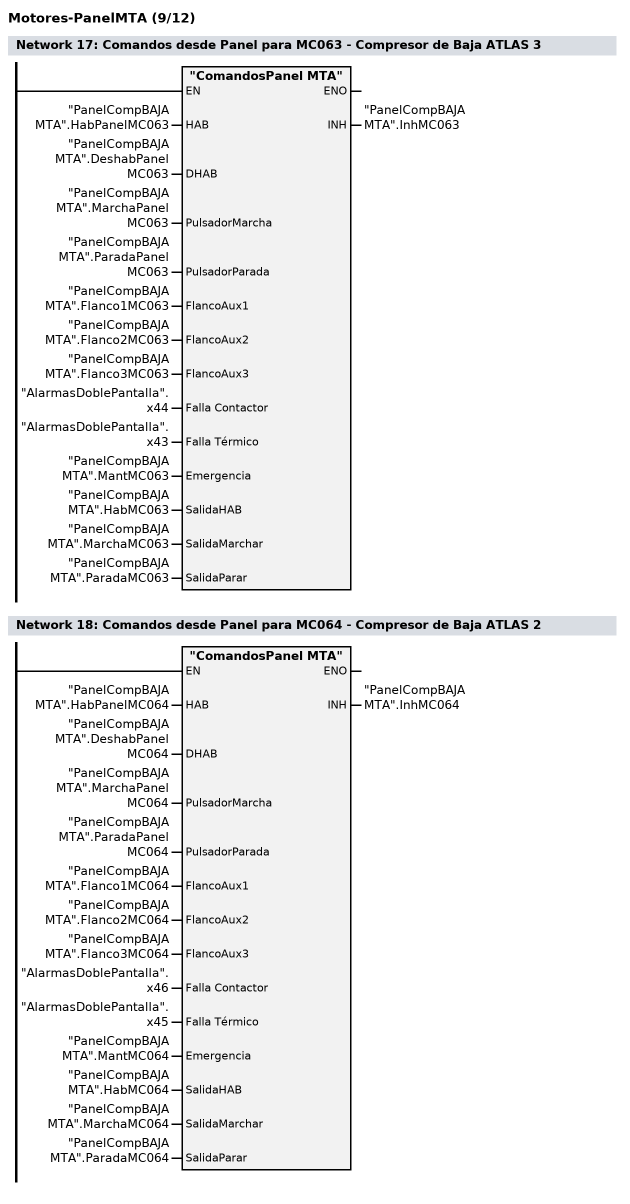
   RUNG wire#powerrail
      "ComandosPanel MTA"(HAB := "PanelCompBAJA MTA".HabPanelMC063, DHAB := "PanelCompBAJA MTA".DeshabPanelMC063, PulsadorMarcha := "PanelCompBAJA MTA".MarchaPanelMC063, PulsadorParada := "PanelCompBAJA MTA".ParadaPanelMC063, FlancoAux1 := "PanelCompBAJA MTA".Flanco1MC063, FlancoAux2 := "PanelCompBAJA MTA".Flanco2MC063, FlancoAux3 := "PanelCompBAJA MTA".Flanco3MC063, "Falla Contactor" := "AlarmasDoblePantalla".x44, "Falla Térmico" := "AlarmasDoblePantalla".x43, Emergencia := "PanelCompBAJA MTA".MantMC063, INH => "PanelCompBAJA MTA".InhMC063, SalidaHAB := "PanelCompBAJA MTA".HabMC063, SalidaMarchar := "PanelCompBAJA MTA".MarchaMC063, SalidaParar := "PanelCompBAJA MTA".ParadaMC063)
   END_RUNG
   // the same network as SCL:
   "ComandosPanel MTA"(HAB := "PanelCompBAJA MTA".HabPanelMC063,
                       DHAB := "PanelCompBAJA MTA".DeshabPanelMC063,
                       PulsadorMarcha := "PanelCompBAJA MTA".MarchaPanelMC063,
                       PulsadorParada := "PanelCompBAJA MTA".ParadaPanelMC063,
                       FlancoAux1 := "PanelCompBAJA MTA".Flanco1MC063,
                       FlancoAux2 := "PanelCompBAJA MTA".Flanco2MC063,
                       FlancoAux3 := "PanelCompBAJA MTA".Flanco3MC063,
                       "Falla Contactor" := "AlarmasDoblePantalla".x44,
                       "Falla Térmico" := "AlarmasDoblePantalla".x43,
                       Emergencia := "PanelCompBAJA MTA".MantMC063,
                       SalidaHAB := "PanelCompBAJA MTA".HabMC063,
                       SalidaMarchar := "PanelCompBAJA MTA".MarchaMC063,
                       SalidaParar := "PanelCompBAJA MTA".ParadaMC063,
                       INH => "PanelCompBAJA MTA".InhMC063);
END_REGION

REGION Network 18: Comandos desde Panel para MC064 - Compresor de Baja ATLAS 2
   RUNG wire#powerrail
      "ComandosPanel MTA"(HAB := "PanelCompBAJA MTA".HabPanelMC064, DHAB := "PanelCompBAJA MTA".DeshabPanelMC064, PulsadorMarcha := "PanelCompBAJA MTA".MarchaPanelMC064, PulsadorParada := "PanelCompBAJA MTA".ParadaPanelMC064, FlancoAux1 := "PanelCompBAJA MTA".Flanco1MC064, FlancoAux2 := "PanelCompBAJA MTA".Flanco2MC064, FlancoAux3 := "PanelCompBAJA MTA".Flanco3MC064, "Falla Contactor" := "AlarmasDoblePantalla".x46, "Falla Térmico" := "AlarmasDoblePantalla".x45, Emergencia := "PanelCompBAJA MTA".MantMC064, INH => "PanelCompBAJA MTA".InhMC064, SalidaHAB := "PanelCompBAJA MTA".HabMC064, SalidaMarchar := "PanelCompBAJA MTA".MarchaMC064, SalidaParar := "PanelCompBAJA MTA".ParadaMC064)
   END_RUNG
   // the same network as SCL:
   "ComandosPanel MTA"(HAB := "PanelCompBAJA MTA".HabPanelMC064,
                       DHAB := "PanelCompBAJA MTA".DeshabPanelMC064,
                       PulsadorMarcha := "PanelCompBAJA MTA".MarchaPanelMC064,
                       PulsadorParada := "PanelCompBAJA MTA".ParadaPanelMC064,
                       FlancoAux1 := "PanelCompBAJA MTA".Flanco1MC064,
                       FlancoAux2 := "PanelCompBAJA MTA".Flanco2MC064,
                       FlancoAux3 := "PanelCompBAJA MTA".Flanco3MC064,
                       "Falla Contactor" := "AlarmasDoblePantalla".x46,
                       "Falla Térmico" := "AlarmasDoblePantalla".x45,
                       Emergencia := "PanelCompBAJA MTA".MantMC064,
                       SalidaHAB := "PanelCompBAJA MTA".HabMC064,
                       SalidaMarchar := "PanelCompBAJA MTA".MarchaMC064,
                       SalidaParar := "PanelCompBAJA MTA".ParadaMC064,
                       INH => "PanelCompBAJA MTA".InhMC064);
END_REGION

REGION Network 19: Comandos desde Panel para MS050 - Secador de Alta ABC1
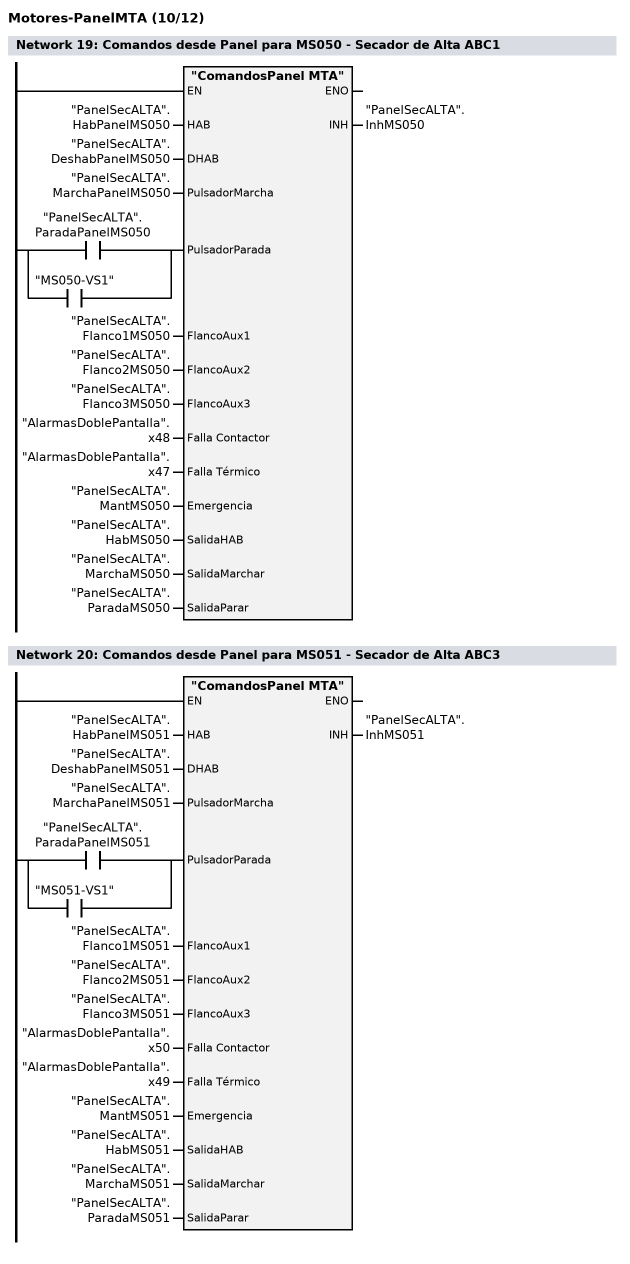
   RUNG wire#powerrail
      "ComandosPanel MTA"(HAB := "PanelSecALTA".HabPanelMS050, DHAB := "PanelSecALTA".DeshabPanelMS050, PulsadorMarcha := "PanelSecALTA".MarchaPanelMS050, PulsadorParada := wire#w1, FlancoAux1 := "PanelSecALTA".Flanco1MS050, FlancoAux2 := "PanelSecALTA".Flanco2MS050, FlancoAux3 := "PanelSecALTA".Flanco3MS050, "Falla Contactor" := "AlarmasDoblePantalla".x48, "Falla Térmico" := "AlarmasDoblePantalla".x47, Emergencia := "PanelSecALTA".MantMS050, INH => "PanelSecALTA".InhMS050, SalidaHAB := "PanelSecALTA".HabMS050, SalidaMarchar := "PanelSecALTA".MarchaMS050, SalidaParar := "PanelSecALTA".ParadaMS050)
   END_RUNG
   RUNG wire#powerrail
      Contact( "PanelSecALTA".ParadaPanelMS050 )
   END_RUNG wire#w1
   RUNG wire#powerrail
      Contact( "MS050-VS1" )
   END_RUNG wire#w1
   // the same network as SCL:
   "ComandosPanel MTA"(HAB := "PanelSecALTA".HabPanelMS050,
                       DHAB := "PanelSecALTA".DeshabPanelMS050,
                       PulsadorMarcha := "PanelSecALTA".MarchaPanelMS050,
                       PulsadorParada := "PanelSecALTA".ParadaPanelMS050 OR "MS050-VS1",
                       FlancoAux1 := "PanelSecALTA".Flanco1MS050,
                       FlancoAux2 := "PanelSecALTA".Flanco2MS050,
                       FlancoAux3 := "PanelSecALTA".Flanco3MS050,
                       "Falla Contactor" := "AlarmasDoblePantalla".x48,
                       "Falla Térmico" := "AlarmasDoblePantalla".x47,
                       Emergencia := "PanelSecALTA".MantMS050,
                       SalidaHAB := "PanelSecALTA".HabMS050,
                       SalidaMarchar := "PanelSecALTA".MarchaMS050,
                       SalidaParar := "PanelSecALTA".ParadaMS050,
                       INH => "PanelSecALTA".InhMS050);
END_REGION

REGION Network 20: Comandos desde Panel para MS051 - Secador de Alta ABC3
   RUNG wire#powerrail
      "ComandosPanel MTA"(HAB := "PanelSecALTA".HabPanelMS051, DHAB := "PanelSecALTA".DeshabPanelMS051, PulsadorMarcha := "PanelSecALTA".MarchaPanelMS051, PulsadorParada := wire#w1, FlancoAux1 := "PanelSecALTA".Flanco1MS051, FlancoAux2 := "PanelSecALTA".Flanco2MS051, FlancoAux3 := "PanelSecALTA".Flanco3MS051, "Falla Contactor" := "AlarmasDoblePantalla".x50, "Falla Térmico" := "AlarmasDoblePantalla".x49, Emergencia := "PanelSecALTA".MantMS051, INH => "PanelSecALTA".InhMS051, SalidaHAB := "PanelSecALTA".HabMS051, SalidaMarchar := "PanelSecALTA".MarchaMS051, SalidaParar := "PanelSecALTA".ParadaMS051)
   END_RUNG
   RUNG wire#powerrail
      Contact( "PanelSecALTA".ParadaPanelMS051 )
   END_RUNG wire#w1
   RUNG wire#powerrail
      Contact( "MS051-VS1" )
   END_RUNG wire#w1
   // the same network as SCL:
   "ComandosPanel MTA"(HAB := "PanelSecALTA".HabPanelMS051,
                       DHAB := "PanelSecALTA".DeshabPanelMS051,
                       PulsadorMarcha := "PanelSecALTA".MarchaPanelMS051,
                       PulsadorParada := "PanelSecALTA".ParadaPanelMS051 OR "MS051-VS1",
                       FlancoAux1 := "PanelSecALTA".Flanco1MS051,
                       FlancoAux2 := "PanelSecALTA".Flanco2MS051,
                       FlancoAux3 := "PanelSecALTA".Flanco3MS051,
                       "Falla Contactor" := "AlarmasDoblePantalla".x50,
                       "Falla Térmico" := "AlarmasDoblePantalla".x49,
                       Emergencia := "PanelSecALTA".MantMS051,
                       SalidaHAB := "PanelSecALTA".HabMS051,
                       SalidaMarchar := "PanelSecALTA".MarchaMS051,
                       SalidaParar := "PanelSecALTA".ParadaMS051,
                       INH => "PanelSecALTA".InhMS051);
END_REGION

REGION Network 21: Comandos desde Panel para MS052 - Secador de Alta ABC2
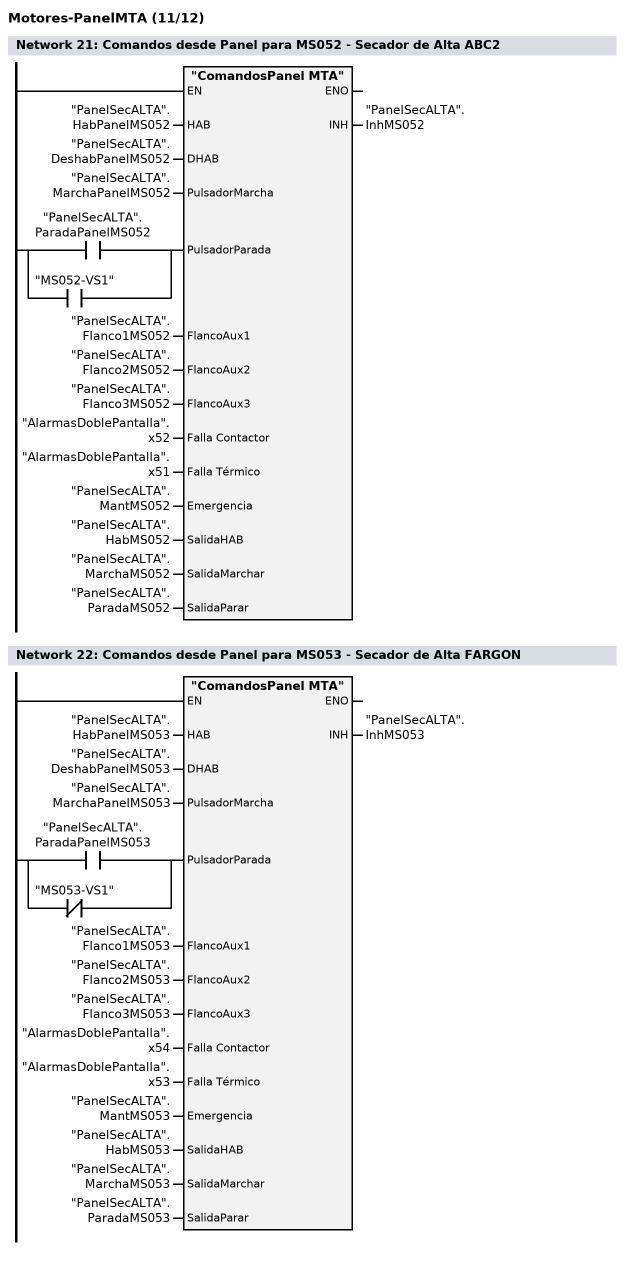
   RUNG wire#powerrail
      "ComandosPanel MTA"(HAB := "PanelSecALTA".HabPanelMS052, DHAB := "PanelSecALTA".DeshabPanelMS052, PulsadorMarcha := "PanelSecALTA".MarchaPanelMS052, PulsadorParada := wire#w1, FlancoAux1 := "PanelSecALTA".Flanco1MS052, FlancoAux2 := "PanelSecALTA".Flanco2MS052, FlancoAux3 := "PanelSecALTA".Flanco3MS052, "Falla Contactor" := "AlarmasDoblePantalla".x52, "Falla Térmico" := "AlarmasDoblePantalla".x51, Emergencia := "PanelSecALTA".MantMS052, INH => "PanelSecALTA".InhMS052, SalidaHAB := "PanelSecALTA".HabMS052, SalidaMarchar := "PanelSecALTA".MarchaMS052, SalidaParar := "PanelSecALTA".ParadaMS052)
   END_RUNG
   RUNG wire#powerrail
      Contact( "PanelSecALTA".ParadaPanelMS052 )
   END_RUNG wire#w1
   RUNG wire#powerrail
      Contact( "MS052-VS1" )
   END_RUNG wire#w1
   // the same network as SCL:
   "ComandosPanel MTA"(HAB := "PanelSecALTA".HabPanelMS052,
                       DHAB := "PanelSecALTA".DeshabPanelMS052,
                       PulsadorMarcha := "PanelSecALTA".MarchaPanelMS052,
                       PulsadorParada := "PanelSecALTA".ParadaPanelMS052 OR "MS052-VS1",
                       FlancoAux1 := "PanelSecALTA".Flanco1MS052,
                       FlancoAux2 := "PanelSecALTA".Flanco2MS052,
                       FlancoAux3 := "PanelSecALTA".Flanco3MS052,
                       "Falla Contactor" := "AlarmasDoblePantalla".x52,
                       "Falla Térmico" := "AlarmasDoblePantalla".x51,
                       Emergencia := "PanelSecALTA".MantMS052,
                       SalidaHAB := "PanelSecALTA".HabMS052,
                       SalidaMarchar := "PanelSecALTA".MarchaMS052,
                       SalidaParar := "PanelSecALTA".ParadaMS052,
                       INH => "PanelSecALTA".InhMS052);
END_REGION

REGION Network 22: Comandos desde Panel para MS053 - Secador de Alta FARGON
   RUNG wire#powerrail
      "ComandosPanel MTA"(HAB := "PanelSecALTA".HabPanelMS053, DHAB := "PanelSecALTA".DeshabPanelMS053, PulsadorMarcha := "PanelSecALTA".MarchaPanelMS053, PulsadorParada := wire#w1, FlancoAux1 := "PanelSecALTA".Flanco1MS053, FlancoAux2 := "PanelSecALTA".Flanco2MS053, FlancoAux3 := "PanelSecALTA".Flanco3MS053, "Falla Contactor" := "AlarmasDoblePantalla".x54, "Falla Térmico" := "AlarmasDoblePantalla".x53, Emergencia := "PanelSecALTA".MantMS053, INH => "PanelSecALTA".InhMS053, SalidaHAB := "PanelSecALTA".HabMS053, SalidaMarchar := "PanelSecALTA".MarchaMS053, SalidaParar := "PanelSecALTA".ParadaMS053)
   END_RUNG
   RUNG wire#powerrail
      Contact( "PanelSecALTA".ParadaPanelMS053 )
   END_RUNG wire#w1
   RUNG wire#powerrail
      I_Contact( "MS053-VS1" )
   END_RUNG wire#w1
   // the same network as SCL:
   "ComandosPanel MTA"(HAB := "PanelSecALTA".HabPanelMS053,
                       DHAB := "PanelSecALTA".DeshabPanelMS053,
                       PulsadorMarcha := "PanelSecALTA".MarchaPanelMS053,
                       PulsadorParada := "PanelSecALTA".ParadaPanelMS053 OR NOT "MS053-VS1",
                       FlancoAux1 := "PanelSecALTA".Flanco1MS053,
                       FlancoAux2 := "PanelSecALTA".Flanco2MS053,
                       FlancoAux3 := "PanelSecALTA".Flanco3MS053,
                       "Falla Contactor" := "AlarmasDoblePantalla".x54,
                       "Falla Térmico" := "AlarmasDoblePantalla".x53,
                       Emergencia := "PanelSecALTA".MantMS053,
                       SalidaHAB := "PanelSecALTA".HabMS053,
                       SalidaMarchar := "PanelSecALTA".MarchaMS053,
                       SalidaParar := "PanelSecALTA".ParadaMS053,
                       INH => "PanelSecALTA".InhMS053);
END_REGION

REGION Network 23: Comandos desde Panel para MS054 - Secador de Baja SULLAIR 1
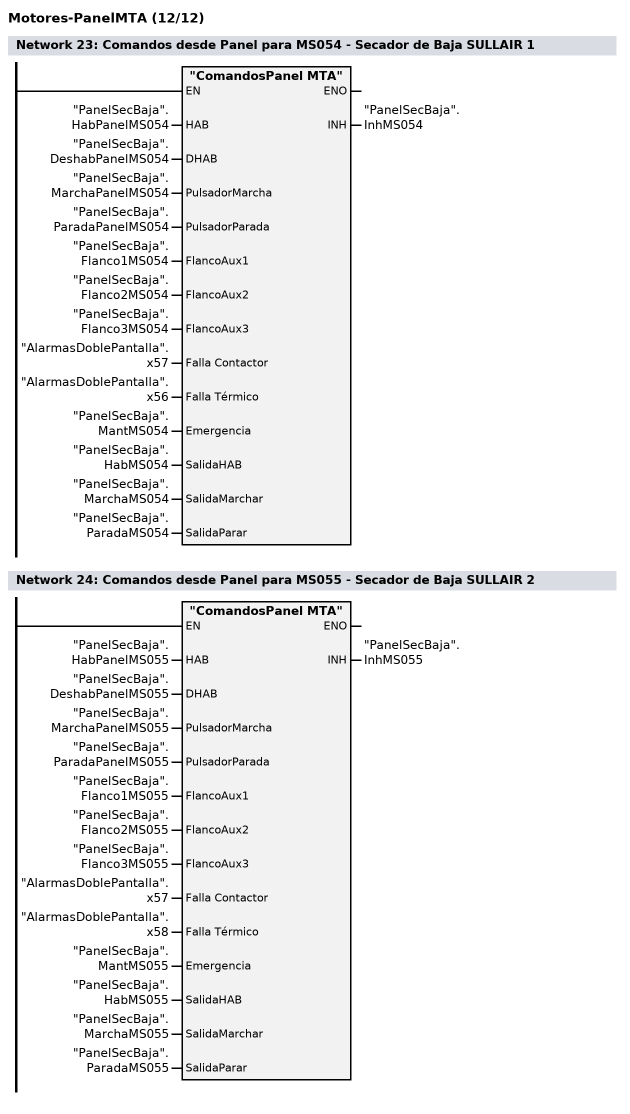
   RUNG wire#powerrail
      "ComandosPanel MTA"(HAB := "PanelSecBaja".HabPanelMS054, DHAB := "PanelSecBaja".DeshabPanelMS054, PulsadorMarcha := "PanelSecBaja".MarchaPanelMS054, PulsadorParada := "PanelSecBaja".ParadaPanelMS054, FlancoAux1 := "PanelSecBaja".Flanco1MS054, FlancoAux2 := "PanelSecBaja".Flanco2MS054, FlancoAux3 := "PanelSecBaja".Flanco3MS054, "Falla Contactor" := "AlarmasDoblePantalla".x57, "Falla Térmico" := "AlarmasDoblePantalla".x56, Emergencia := "PanelSecBaja".MantMS054, INH => "PanelSecBaja".InhMS054, SalidaHAB := "PanelSecBaja".HabMS054, SalidaMarchar := "PanelSecBaja".MarchaMS054, SalidaParar := "PanelSecBaja".ParadaMS054)
   END_RUNG
   // the same network as SCL:
   "ComandosPanel MTA"(HAB := "PanelSecBaja".HabPanelMS054,
                       DHAB := "PanelSecBaja".DeshabPanelMS054,
                       PulsadorMarcha := "PanelSecBaja".MarchaPanelMS054,
                       PulsadorParada := "PanelSecBaja".ParadaPanelMS054,
                       FlancoAux1 := "PanelSecBaja".Flanco1MS054,
                       FlancoAux2 := "PanelSecBaja".Flanco2MS054,
                       FlancoAux3 := "PanelSecBaja".Flanco3MS054,
                       "Falla Contactor" := "AlarmasDoblePantalla".x57,
                       "Falla Térmico" := "AlarmasDoblePantalla".x56,
                       Emergencia := "PanelSecBaja".MantMS054,
                       SalidaHAB := "PanelSecBaja".HabMS054,
                       SalidaMarchar := "PanelSecBaja".MarchaMS054,
                       SalidaParar := "PanelSecBaja".ParadaMS054,
                       INH => "PanelSecBaja".InhMS054);
END_REGION

REGION Network 24: Comandos desde Panel para MS055 - Secador de Baja SULLAIR 2
   RUNG wire#powerrail
      "ComandosPanel MTA"(HAB := "PanelSecBaja".HabPanelMS055, DHAB := "PanelSecBaja".DeshabPanelMS055, PulsadorMarcha := "PanelSecBaja".MarchaPanelMS055, PulsadorParada := "PanelSecBaja".ParadaPanelMS055, FlancoAux1 := "PanelSecBaja".Flanco1MS055, FlancoAux2 := "PanelSecBaja".Flanco2MS055, FlancoAux3 := "PanelSecBaja".Flanco3MS055, "Falla Contactor" := "AlarmasDoblePantalla".x57, "Falla Térmico" := "AlarmasDoblePantalla".x58, Emergencia := "PanelSecBaja".MantMS055, INH => "PanelSecBaja".InhMS055, SalidaHAB := "PanelSecBaja".HabMS055, SalidaMarchar := "PanelSecBaja".MarchaMS055, SalidaParar := "PanelSecBaja".ParadaMS055)
   END_RUNG
   // the same network as SCL:
   "ComandosPanel MTA"(HAB := "PanelSecBaja".HabPanelMS055,
                       DHAB := "PanelSecBaja".DeshabPanelMS055,
                       PulsadorMarcha := "PanelSecBaja".MarchaPanelMS055,
                       PulsadorParada := "PanelSecBaja".ParadaPanelMS055,
                       FlancoAux1 := "PanelSecBaja".Flanco1MS055,
                       FlancoAux2 := "PanelSecBaja".Flanco2MS055,
                       FlancoAux3 := "PanelSecBaja".Flanco3MS055,
                       "Falla Contactor" := "AlarmasDoblePantalla".x57,
                       "Falla Térmico" := "AlarmasDoblePantalla".x58,
                       Emergencia := "PanelSecBaja".MantMS055,
                       SalidaHAB := "PanelSecBaja".HabMS055,
                       SalidaMarchar := "PanelSecBaja".MarchaMS055,
                       SalidaParar := "PanelSecBaja".ParadaMS055,
                       INH => "PanelSecBaja".InhMS055);
END_REGION
END_FUNCTION

FUNCTION "ComandosPanel MTA" : Void   // FC19, LAD
{ S7_Optimized_Access := 'FALSE' }
VERSION : 0.1
   VAR_TEMP   // added for the SCL form of the ladder/FBD networks
      _w1 : Bool;
   END_VAR
BEGIN

REGION Network 1
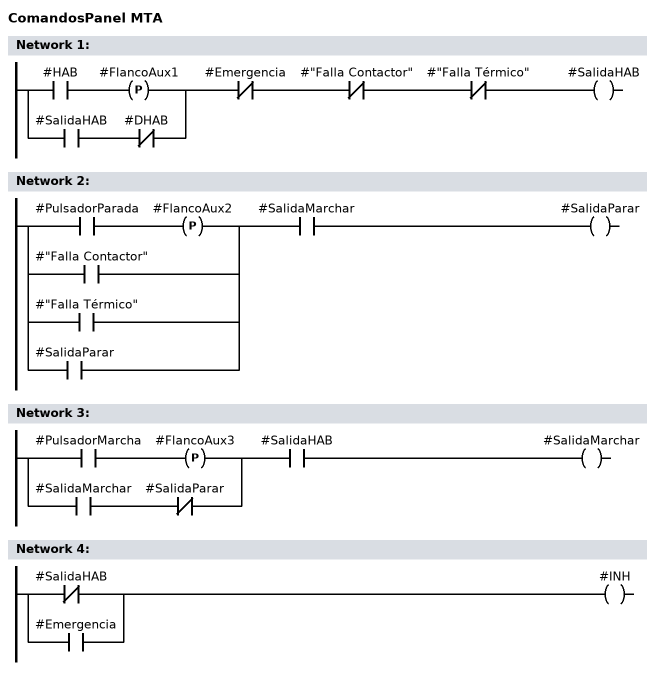
   RUNG wire#powerrail
      Contact( #HAB )
      P_Trig( #FlancoAux1 )
      wire#w1
      I_Contact( #Emergencia )
      I_Contact( #"Falla Contactor" )
      I_Contact( #"Falla Térmico" )
      Coil( #SalidaHAB )
   END_RUNG
   RUNG wire#powerrail
      Contact( #SalidaHAB )
      I_Contact( #DHAB )
   END_RUNG wire#w1
   // the same network as SCL:
   #_w1 := #HAB AND NOT #FlancoAux1;   // rising edge
   #FlancoAux1 := #HAB;
   #SalidaHAB := (#_w1 OR (#SalidaHAB AND NOT #DHAB)) AND NOT #Emergencia AND NOT #"Falla Contactor" AND NOT #"Falla Térmico";
END_REGION

REGION Network 2
   RUNG wire#powerrail
      Contact( #PulsadorParada )
      P_Trig( #FlancoAux2 )
      wire#w1
      Contact( #SalidaMarchar )
      Coil( #SalidaParar )
   END_RUNG
   RUNG wire#powerrail
      Contact( #"Falla Contactor" )
   END_RUNG wire#w1
   RUNG wire#powerrail
      Contact( #"Falla Térmico" )
   END_RUNG wire#w1
   RUNG wire#powerrail
      Contact( #SalidaParar )
   END_RUNG wire#w1
   // the same network as SCL:
   #_w1 := #PulsadorParada AND NOT #FlancoAux2;   // rising edge
   #FlancoAux2 := #PulsadorParada;
   #SalidaParar := (#_w1 OR #"Falla Contactor" OR #"Falla Térmico" OR #SalidaParar) AND #SalidaMarchar;
END_REGION

REGION Network 3
   RUNG wire#powerrail
      Contact( #PulsadorMarcha )
      P_Trig( #FlancoAux3 )
      wire#w1
      Contact( #SalidaHAB )
      Coil( #SalidaMarchar )
   END_RUNG
   RUNG wire#powerrail
      Contact( #SalidaMarchar )
      I_Contact( #SalidaParar )
   END_RUNG wire#w1
   // the same network as SCL:
   #_w1 := #PulsadorMarcha AND NOT #FlancoAux3;   // rising edge
   #FlancoAux3 := #PulsadorMarcha;
   #SalidaMarchar := (#_w1 OR (#SalidaMarchar AND NOT #SalidaParar)) AND #SalidaHAB;
END_REGION

REGION Network 4
   RUNG wire#powerrail
      I_Contact( #SalidaHAB )
      wire#w1
      Coil( #INH )
   END_RUNG
   RUNG wire#powerrail
      Contact( #Emergencia )
   END_RUNG wire#w1
   // the same network as SCL:
   #INH := NOT #SalidaHAB OR #Emergencia;
END_REGION
END_FUNCTION

FUNCTION "FC-ANIM-CMP" : Void   // FC43, LAD
{ S7_Optimized_Access := 'FALSE' }
VERSION : 0.1
BEGIN

REGION Network 1
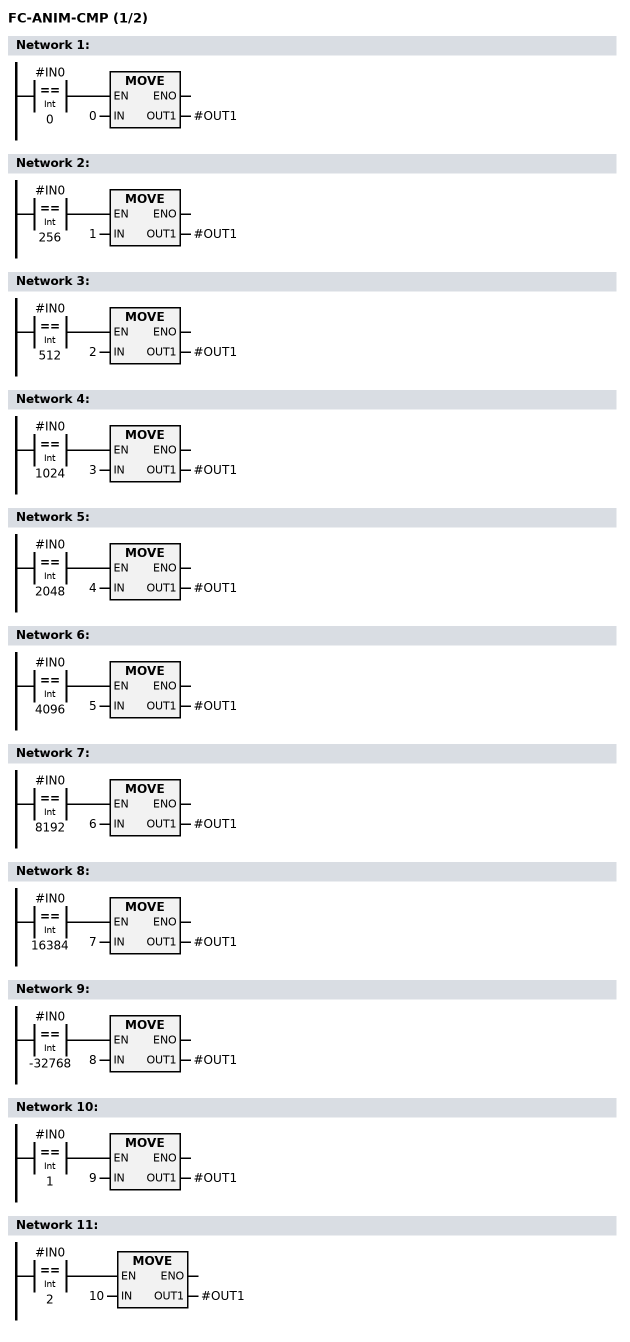
   RUNG wire#powerrail
      { S7_Templates := "SrcType := Int" } EQ_Contact(in1 := #IN0, in2 := 0)
      { S7_GenerateENO := "TRUE" } Move(in := 0, out1 => #OUT1)
   END_RUNG
   // the same network as SCL:
   IF #IN0 = 0 THEN #OUT1 := 0; END_IF;
END_REGION

REGION Network 2
   RUNG wire#powerrail
      { S7_Templates := "SrcType := Int" } EQ_Contact(in1 := #IN0, in2 := 256)
      { S7_GenerateENO := "TRUE" } Move(in := 1, out1 => #OUT1)
   END_RUNG
   // the same network as SCL:
   IF #IN0 = 256 THEN #OUT1 := 1; END_IF;
END_REGION

REGION Network 3
   RUNG wire#powerrail
      { S7_Templates := "SrcType := Int" } EQ_Contact(in1 := #IN0, in2 := 512)
      { S7_GenerateENO := "TRUE" } Move(in := 2, out1 => #OUT1)
   END_RUNG
   // the same network as SCL:
   IF #IN0 = 512 THEN #OUT1 := 2; END_IF;
END_REGION

REGION Network 4
   RUNG wire#powerrail
      { S7_Templates := "SrcType := Int" } EQ_Contact(in1 := #IN0, in2 := 1024)
      { S7_GenerateENO := "TRUE" } Move(in := 3, out1 => #OUT1)
   END_RUNG
   // the same network as SCL:
   IF #IN0 = 1024 THEN #OUT1 := 3; END_IF;
END_REGION

REGION Network 5
   RUNG wire#powerrail
      { S7_Templates := "SrcType := Int" } EQ_Contact(in1 := #IN0, in2 := 2048)
      { S7_GenerateENO := "TRUE" } Move(in := 4, out1 => #OUT1)
   END_RUNG
   // the same network as SCL:
   IF #IN0 = 2048 THEN #OUT1 := 4; END_IF;
END_REGION

REGION Network 6
   RUNG wire#powerrail
      { S7_Templates := "SrcType := Int" } EQ_Contact(in1 := #IN0, in2 := 4096)
      { S7_GenerateENO := "TRUE" } Move(in := 5, out1 => #OUT1)
   END_RUNG
   // the same network as SCL:
   IF #IN0 = 4096 THEN #OUT1 := 5; END_IF;
END_REGION

REGION Network 7
   RUNG wire#powerrail
      { S7_Templates := "SrcType := Int" } EQ_Contact(in1 := #IN0, in2 := 8192)
      { S7_GenerateENO := "TRUE" } Move(in := 6, out1 => #OUT1)
   END_RUNG
   // the same network as SCL:
   IF #IN0 = 8192 THEN #OUT1 := 6; END_IF;
END_REGION

REGION Network 8
   RUNG wire#powerrail
      { S7_Templates := "SrcType := Int" } EQ_Contact(in1 := #IN0, in2 := 16384)
      { S7_GenerateENO := "TRUE" } Move(in := 7, out1 => #OUT1)
   END_RUNG
   // the same network as SCL:
   IF #IN0 = 16384 THEN #OUT1 := 7; END_IF;
END_REGION

REGION Network 9
   RUNG wire#powerrail
      { S7_Templates := "SrcType := Int" } EQ_Contact(in1 := #IN0, in2 := -32768)
      { S7_GenerateENO := "TRUE" } Move(in := 8, out1 => #OUT1)
   END_RUNG
   // the same network as SCL:
   IF #IN0 = (-32768) THEN #OUT1 := 8; END_IF;
END_REGION

REGION Network 10
   RUNG wire#powerrail
      { S7_Templates := "SrcType := Int" } EQ_Contact(in1 := #IN0, in2 := 1)
      { S7_GenerateENO := "TRUE" } Move(in := 9, out1 => #OUT1)
   END_RUNG
   // the same network as SCL:
   IF #IN0 = 1 THEN #OUT1 := 9; END_IF;
END_REGION

REGION Network 11
   RUNG wire#powerrail
      { S7_Templates := "SrcType := Int" } EQ_Contact(in1 := #IN0, in2 := 2)
      { S7_GenerateENO := "TRUE" } Move(in := 10, out1 => #OUT1)
   END_RUNG
   // the same network as SCL:
   IF #IN0 = 2 THEN #OUT1 := 10; END_IF;
END_REGION

REGION Network 12
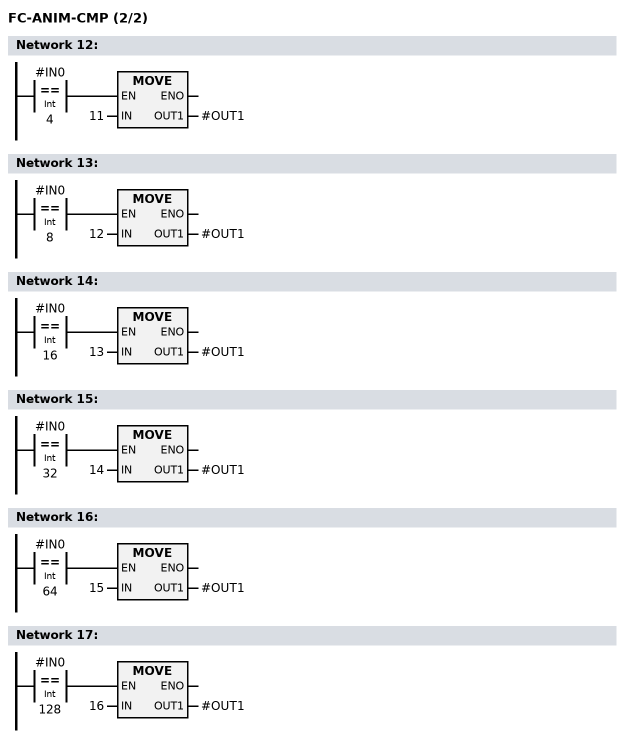
   RUNG wire#powerrail
      { S7_Templates := "SrcType := Int" } EQ_Contact(in1 := #IN0, in2 := 4)
      { S7_GenerateENO := "TRUE" } Move(in := 11, out1 => #OUT1)
   END_RUNG
   // the same network as SCL:
   IF #IN0 = 4 THEN #OUT1 := 11; END_IF;
END_REGION

REGION Network 13
   RUNG wire#powerrail
      { S7_Templates := "SrcType := Int" } EQ_Contact(in1 := #IN0, in2 := 8)
      { S7_GenerateENO := "TRUE" } Move(in := 12, out1 => #OUT1)
   END_RUNG
   // the same network as SCL:
   IF #IN0 = 8 THEN #OUT1 := 12; END_IF;
END_REGION

REGION Network 14
   RUNG wire#powerrail
      { S7_Templates := "SrcType := Int" } EQ_Contact(in1 := #IN0, in2 := 16)
      { S7_GenerateENO := "TRUE" } Move(in := 13, out1 => #OUT1)
   END_RUNG
   // the same network as SCL:
   IF #IN0 = 16 THEN #OUT1 := 13; END_IF;
END_REGION

REGION Network 15
   RUNG wire#powerrail
      { S7_Templates := "SrcType := Int" } EQ_Contact(in1 := #IN0, in2 := 32)
      { S7_GenerateENO := "TRUE" } Move(in := 14, out1 => #OUT1)
   END_RUNG
   // the same network as SCL:
   IF #IN0 = 32 THEN #OUT1 := 14; END_IF;
END_REGION

REGION Network 16
   RUNG wire#powerrail
      { S7_Templates := "SrcType := Int" } EQ_Contact(in1 := #IN0, in2 := 64)
      { S7_GenerateENO := "TRUE" } Move(in := 15, out1 => #OUT1)
   END_RUNG
   // the same network as SCL:
   IF #IN0 = 64 THEN #OUT1 := 15; END_IF;
END_REGION

REGION Network 17
   RUNG wire#powerrail
      { S7_Templates := "SrcType := Int" } EQ_Contact(in1 := #IN0, in2 := 128)
      { S7_GenerateENO := "TRUE" } Move(in := 16, out1 => #OUT1)
   END_RUNG
   // the same network as SCL:
   IF #IN0 = 128 THEN #OUT1 := 16; END_IF;
END_REGION
END_FUNCTION

// folder: Panel/Iluminación

FUNCTION "IluminaciónMTA" : Void   // FC23, LAD
{ S7_Optimized_Access := 'FALSE' }
VERSION : 0.1
// LUC - 05/08/2020
   VAR_TEMP   // added for the SCL form of the ladder/FBD networks
      _s5time1 : S5Time;
   END_VAR
BEGIN

REGION Network 1: Seteo de temporizador desde panel
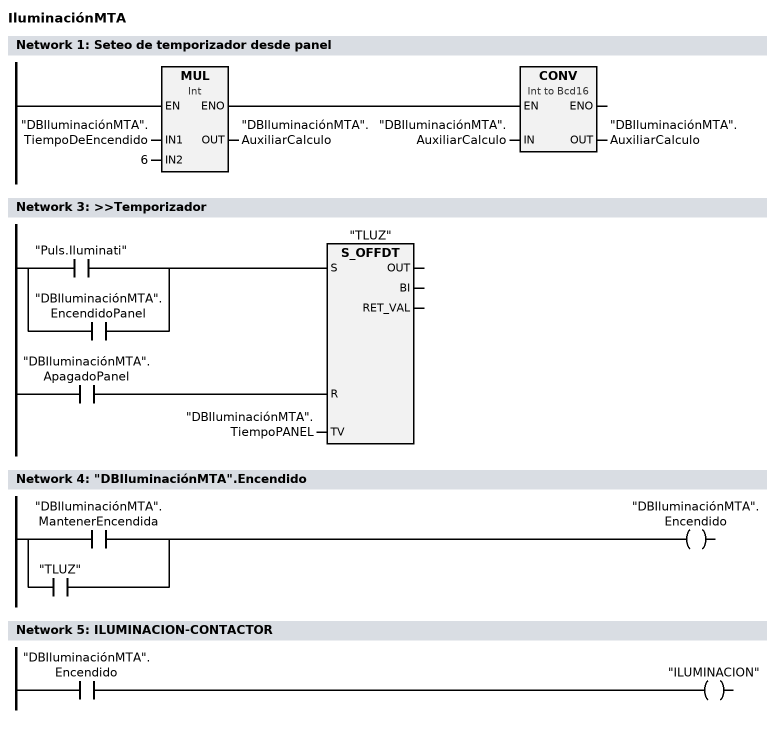
   RUNG wire#powerrail
      { S7_Templates := "SrcType := Int"; S7_GenerateENO := "TRUE" } Mul(in1 := "DBIluminaciónMTA".TiempoDeEncendido, in2 := 6, out => "DBIluminaciónMTA".AuxiliarCalculo)
      { S7_Templates := "[SrcType := Int, DestType := Bcd16]"; S7_GenerateENO := "TRUE" } Convert(in := "DBIluminaciónMTA".AuxiliarCalculo, out => "DBIluminaciónMTA".AuxiliarCalculo)
   END_RUNG
   // the same network as SCL:
   // ENO of a box is taken as its EN; it also drops when the box reports an error
   "DBIluminaciónMTA".AuxiliarCalculo := "DBIluminaciónMTA".TiempoDeEncendido * 6;
   "DBIluminaciónMTA".AuxiliarCalculo := INT_TO_BCD16("DBIluminaciónMTA".AuxiliarCalculo);
END_REGION

REGION Network 2 (STL): Seteo de temporizador desde panel
         L     12288;
         L     "DBIluminaciónMTA".AuxiliarCalculo;
         OW;
         T     "DBIluminaciónMTA".TiempoPANEL;
         NOP   0;
END_REGION

REGION Network 3: >>Temporizador
   RUNG wire#powerrail
      Contact( "Puls.Iluminati" )
      wire#w1
      S_OFFDT(T_NO := "TLUZ", R := wire#w2, TV := "DBIluminaciónMTA".TiempoPANEL, BI =>, RET_VAL =>)
   END_RUNG
   RUNG wire#powerrail
      Contact( "DBIluminaciónMTA".EncendidoPanel )
   END_RUNG wire#w1
   RUNG wire#powerrail
      Contact( "DBIluminaciónMTA".ApagadoPanel )
   END_RUNG wire#w2
   // the same network as SCL:
   #_s5time1 := S_OFFDT(T_NO := "TLUZ",
                        S := "Puls.Iluminati" OR "DBIluminaciónMTA".EncendidoPanel,
                        R := "DBIluminaciónMTA".ApagadoPanel,
                        TV := "DBIluminaciónMTA".TiempoPANEL);
END_REGION

REGION Network 4: "DBIluminaciónMTA".Encendido
   RUNG wire#powerrail
      Contact( "DBIluminaciónMTA".MantenerEncendida )
      wire#w1
      Coil( "DBIluminaciónMTA".Encendido )
   END_RUNG
   RUNG wire#powerrail
      Contact( "TLUZ" )
   END_RUNG wire#w1
   // the same network as SCL:
   "DBIluminaciónMTA".Encendido := "DBIluminaciónMTA".MantenerEncendida OR "TLUZ";
END_REGION

REGION Network 5: ILUMINACION-CONTACTOR
   RUNG wire#powerrail
      Contact( "DBIluminaciónMTA".Encendido )
      Coil( "ILUMINACION" )
   END_RUNG
   // the same network as SCL:
   "ILUMINACION" := "DBIluminaciónMTA".Encendido;
END_REGION
END_FUNCTION

// folder: Secadores/Alta

FUNCTION "EnclavSecAltaMTA" : Void   // FC12, LAD
{ S7_Optimized_Access := 'FALSE' }
VERSION : 0.1
BEGIN

REGION Network 1: Arranque automático MS050
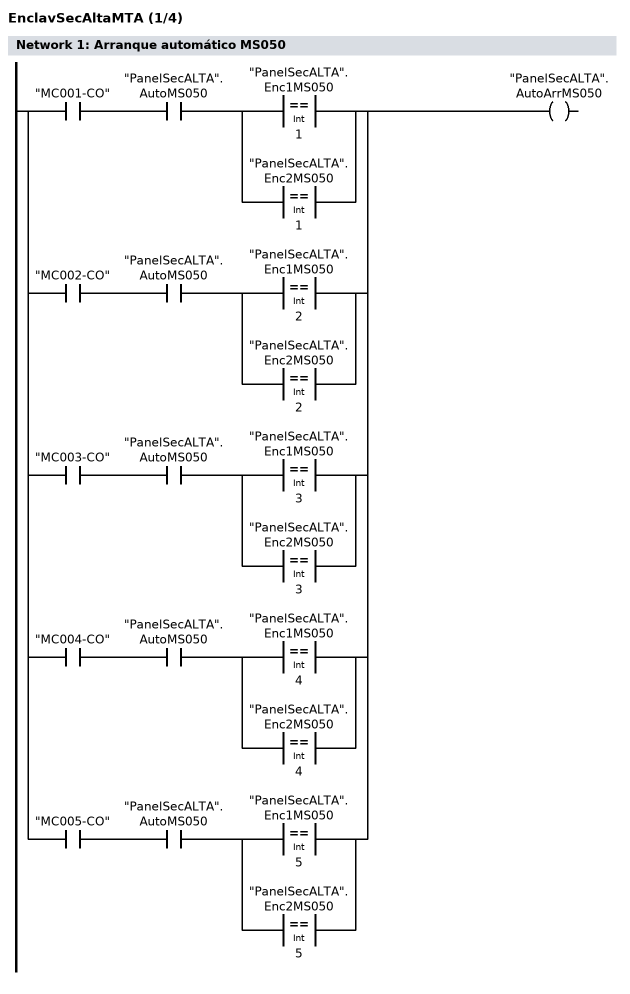
   "PanelSecALTA".AutoArrMS050 := ("MC001-CO" AND "PanelSecALTA".AutoMS050 AND (("PanelSecALTA".Enc1MS050 = 1) OR ("PanelSecALTA".Enc2MS050 = 1))) OR ("MC002-CO" AND "PanelSecALTA".AutoMS050 AND (("PanelSecALTA".Enc1MS050 = 2) OR ("PanelSecALTA".Enc2MS050 = 2))) OR ("MC003-CO" AND "PanelSecALTA".AutoMS050 AND (("PanelSecALTA".Enc1MS050 = 3) OR ("PanelSecALTA".Enc2MS050 = 3))) OR ("MC004-CO" AND "PanelSecALTA".AutoMS050 AND (("PanelSecALTA".Enc1MS050 = 4) OR ("PanelSecALTA".Enc2MS050 = 4))) OR ("MC005-CO" AND "PanelSecALTA".AutoMS050 AND (("PanelSecALTA".Enc1MS050 = 5) OR ("PanelSecALTA".Enc2MS050 = 5)));
END_REGION

REGION Network 2: Arranque automático MS051
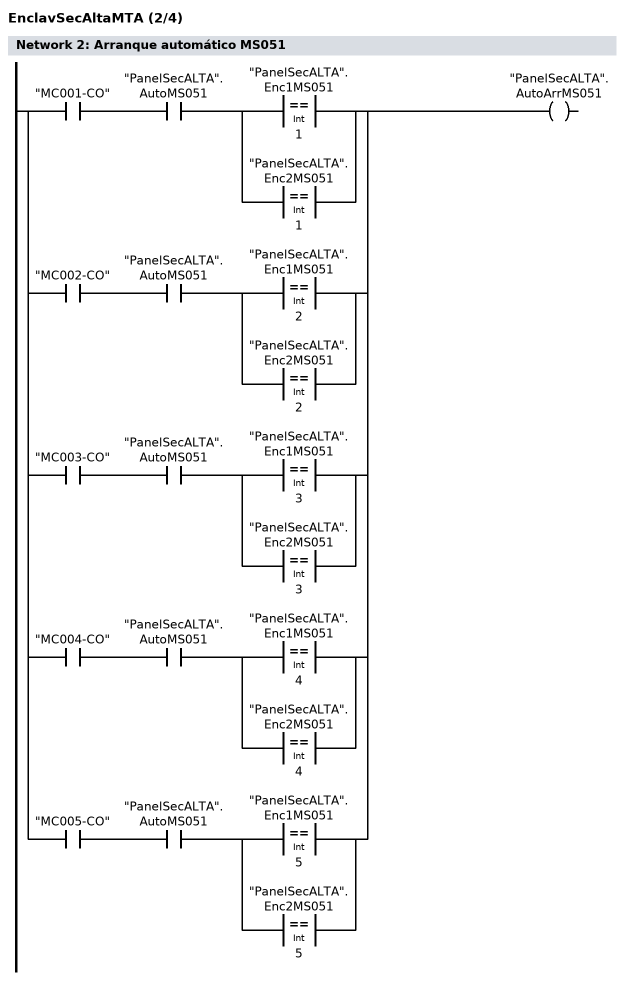
   "PanelSecALTA".AutoArrMS051 := ("MC001-CO" AND "PanelSecALTA".AutoMS051 AND (("PanelSecALTA".Enc1MS051 = 1) OR ("PanelSecALTA".Enc2MS051 = 1))) OR ("MC002-CO" AND "PanelSecALTA".AutoMS051 AND (("PanelSecALTA".Enc1MS051 = 2) OR ("PanelSecALTA".Enc2MS051 = 2))) OR ("MC003-CO" AND "PanelSecALTA".AutoMS051 AND (("PanelSecALTA".Enc1MS051 = 3) OR ("PanelSecALTA".Enc2MS051 = 3))) OR ("MC004-CO" AND "PanelSecALTA".AutoMS051 AND (("PanelSecALTA".Enc1MS051 = 4) OR ("PanelSecALTA".Enc2MS051 = 4))) OR ("MC005-CO" AND "PanelSecALTA".AutoMS051 AND (("PanelSecALTA".Enc1MS051 = 5) OR ("PanelSecALTA".Enc2MS051 = 5)));
END_REGION

REGION Network 3: Arranque automático MS052